// Mitsubishi GX Works2 project: 20国轩1次注液出1031   PLC: Q06UDEH (continued)
  PackCommunication20105 : PackCommunication;
  PackCommunication20106 : PackCommunication;
  PackCommunication20107 : PackCommunication;
  PackCommunication20108 : PackCommunication;
  PackCommunication20109 : PackCommunication;
  PackCommunicationIO20102 : PackCommunicationIO;
  PackCommunicationIO20103 : PackCommunicationIO;
  PackCommunicationIO20104 : PackCommunicationIO;
  PackCommunicationIO20105 : PackCommunicationIO;
  PackCommunicationIO20106 : PackCommunicationIO;
  PackCommunicationIO20107 : PackCommunicationIO;
  PackCommunicationIO20108 : PackCommunicationIO;
  PackCommunicationIO20109 : PackCommunicationIO;
  m_TPU1TaskComplete : TP;  (* U1完成延时 *)
  m_tU1TaskComplete : TIME;  (* U1完成延时 *)
  m_xU1TaskComplete : BOOL;  (* U1完成延时 *)
  m_TPU2TaskComplete : TP;  (* U2完成延时 *)
  m_tU2TaskComplete : TIME;  (* U2完成延时 *)
  m_xU2TaskComplete : BOOL;  (* U2完成延时 *)
  m_TPU3TaskComplete : TP;  (* U3完成延时 *)
  m_tU3TaskComplete : TIME;  (* U3完成延时 *)
  m_xU3TaskComplete : BOOL;  (* U3完成延时 *)
  m_TPU4TaskComplete : TP;  (* U4完成延时 *)
  m_tU4TaskComplete : TIME;  (* U4完成延时 *)
  m_xU4TaskComplete : BOOL;  (* U4完成延时 *)
  m_TonU1TaskStart : TON;  (* U1任务开始延时 *)
  m_tU1TaskStart : TIME;  (* U1任务开始延时 *)
  m_xU1TaskStart : BOOL;  (* U1任务开始延时 *)
  m_TonU2TaskStart : TON;  (* U2任务开始延时 *)
  m_tU2TaskStart : TIME;  (* U2任务开始延时 *)
  m_xU2TaskStart : BOOL;  (* U2任务开始延时 *)
  m_TonU3TaskStart : TON;  (* U3任务开始延时 *)
  m_tU3TaskStart : TIME;  (* U3任务开始延时 *)
  m_xU3TaskStart : BOOL;  (* U3任务开始延时 *)
  m_TonU4TaskStart : TON;  (* U4任务开始延时 *)
  m_tU4TaskStart : TIME;  (* U4任务开始延时 *)
  m_xU4TaskStart : BOOL;  (* U4任务开始延时 *)
  ConveyorIO201221 : ConveyorIO;  (* 虚构的 *)
  Conveyor201221 : Conveyor;  (* 虚构的 *)
  ConveyorIO20119 : ConveyorIO;
  Conveyor20119 : Conveyor;
END_VAR
Conveyor20101(ConveyorMotor:=	ConveyorIO20101);	
(*ConveyorIO20101.xPosLimit:=XA; 	*)
(*ConveyorIO20101.xNegLimit:=X7F; 	*)
ConveyorIO20101.xCWPresent:=X8; 
ConveyorIO20101.xNegLimit:=NOT X9;
(*ConveyorIO20101.xCCWPresent:=X9; 	*)
Y208:=ConveyorIO20101.xMotorCW; 	
Y209:=ConveyorIO20101.xMotorCCW; 	
ConveyorIO20101.xForward:=M500; 	
ConveyorIO20101.xBackward:=M501; 	
M301:= NOT ConveyorIO20101.xEmpty; 	
F401:=ConveyorIO20101.xError; 	
ConveyorIO20101.diDeviceID:=20101; 
ConveyorIO20101.tLoadDelay:=T#2s;	

Conveyor20102(ConveyorMotor:=	ConveyorIO20102);
ConveyorIO20102.xCCWPresent:=X13; 	
Y20A:=ConveyorIO20102.xMotorCW; 	
Y20B:=ConveyorIO20102.xMotorCCW; 	
ConveyorIO20102.xForward:=M502; 	
ConveyorIO20102.xBackward:=M503; 	
M302:= NOT ConveyorIO20102.xEmpty; 	
F402:=ConveyorIO20102.xError; 	
ConveyorIO20102.diDeviceID:=20102;
ConveyorIO20102.tLoadDelay:=T#7s; 
ConveyorIO20102.xloadCCW:=1;	

Conveyor201021(ConveyorMotor:=	ConveyorIO201021);	
ConveyorIO201021.xCWPresent:=X76; 	
M334:= NOT ConveyorIO201021.xEmpty; 	
F434:=ConveyorIO201021.xError; 	
ConveyorIO201021.diDeviceID:=20102; 	
ConveyorIO201021.tLoadDelay:=T#2s;

Conveyor20103(ConveyorMotor:=	ConveyorIO20103);	
ConveyorIO20103.xCCWPresent:=X14; 	
Y20C:=ConveyorIO20103.xMotorCW; 	
Y20D:=ConveyorIO20103.xMotorCCW; 	
ConveyorIO20103.xForward:=M504; 	
ConveyorIO20103.xBackward:=M505; 	
M303:= NOT ConveyorIO20103.xEmpty; 	
F403:=ConveyorIO20103.xError; 	
ConveyorIO20103.diDeviceID:=20103; 
ConveyorIO20103.tLoadDelay:=T#7s; 	
ConveyorIO20103.xloadCCW:=1;	

Conveyor201031(ConveyorMotor:=	ConveyorIO201031);	
ConveyorIO201031.xCWPresent:=X77; 	
M335:= NOT ConveyorIO201031.xEmpty; 	
F435:=ConveyorIO201031.xError; 	
ConveyorIO201031.diDeviceID:=20103; 	
ConveyorIO201031.tLoadDelay:=T#2s;

Conveyor20104(ConveyorMotor:=	ConveyorIO20104);	
ConveyorIO20104.xCCWPresent:=X15; 	
Y20E:=ConveyorIO20104.xMotorCW; 	
Y20F:=ConveyorIO20104.xMotorCCW; 	
ConveyorIO20104.xForward:=M506; 	
ConveyorIO20104.xBackward:=M507; 	
M304:= NOT ConveyorIO20104.xEmpty; 	
F404:=ConveyorIO20104.xError; 	
ConveyorIO20104.diDeviceID:=20104; 
ConveyorIO20104.tLoadDelay:=T#7s; 	
ConveyorIO20104.xloadCCW:=1;		


Conveyor201041(ConveyorMotor:=	ConveyorIO201041);	
ConveyorIO201041.xCWPresent:=X78; 	
M336:= NOT ConveyorIO201041.xEmpty; 	
F436:=ConveyorIO201041.xError; 	
ConveyorIO201041.diDeviceID:=20104; 	
ConveyorIO201041.tLoadDelay:=T#2s;

Conveyor20105(ConveyorMotor:=	ConveyorIO20105);	
ConveyorIO20105.xCCWPresent:=X16; 	
Y210:=ConveyorIO20105.xMotorCW; 	
Y211:=ConveyorIO20105.xMotorCCW; 	
ConveyorIO20105.xForward:=M508; 	
ConveyorIO20105.xBackward:=M509; 	
M305:= NOT ConveyorIO20105.xEmpty; 	
F405:=ConveyorIO20105.xError; 	
ConveyorIO20105.diDeviceID:=20105;		
ConveyorIO20105.tLoadDelay:=T#7s; 	
ConveyorIO20105.xloadCCW:=1;	
				
Conveyor201051(ConveyorMotor:=	ConveyorIO201051);	
ConveyorIO201051.xCWPresent:=X79; 	
M337:= NOT ConveyorIO201051.xEmpty; 	
F437:=ConveyorIO201051.xError; 	
ConveyorIO201051.diDeviceID:=20105; 	
ConveyorIO201051.tLoadDelay:=T#2s;

Conveyor20106(ConveyorMotor:=	ConveyorIO20106);	(*电池X9C*)
ConveyorIO20106.xCCWPresent:=X18; 	
Y212:=ConveyorIO20106.xMotorCW; 	
Y213:=ConveyorIO20106.xMotorCCW; 	
ConveyorIO20106.xForward:=M510; 	
ConveyorIO20106.xBackward:=M511; 	
M306:= NOT ConveyorIO20106.xEmpty; 	
F406:=ConveyorIO20106.xError; 	
ConveyorIO20106.diDeviceID:=20106; 
ConveyorIO20106.tLoadDelay:=T#7s;
ConveyorIO20106.xloadCCW:=1;	 		

Conveyor201061(ConveyorMotor:=	ConveyorIO201061);	
ConveyorIO201061.xCWPresent:=X7A; 	
M338:= NOT ConveyorIO201061.xEmpty; 	
F438:=ConveyorIO201061.xError; 	
ConveyorIO201061.diDeviceID:=20106;
ConveyorIO201061.tLoadDelay:=T#2s; 	

Conveyor20107(ConveyorMotor:=	ConveyorIO20107);	(*电池X9D*)
ConveyorIO20107.xCCWPresent:=X19; 	
Y214:=ConveyorIO20107.xMotorCW; 	
Y215:=ConveyorIO20107.xMotorCCW; 	
ConveyorIO20107.xForward:=M512; 	
ConveyorIO20107.xBackward:=M513; 	
M307:= NOT ConveyorIO20107.xEmpty; 	
F407:=ConveyorIO20107.xError; 	
ConveyorIO20107.diDeviceID:=20107; 
ConveyorIO20107.tLoadDelay:=T#7s; 	
ConveyorIO20107.xloadCCW:=1;	

Conveyor201071(ConveyorMotor:=	ConveyorIO201071);	
ConveyorIO201071.xCWPresent:=X7B; 	
M339:= NOT ConveyorIO201071.xEmpty; 	
F439:=ConveyorIO201071.xError; 	
ConveyorIO201071.diDeviceID:=20107; 	
ConveyorIO201071.tLoadDelay:=T#2s;

Conveyor20108(ConveyorMotor:=	ConveyorIO20108);	(*电池x9e*)
ConveyorIO20108.xCCWPresent:=X1A; 	
Y216:=ConveyorIO20108.xMotorCW; 	
Y217:=ConveyorIO20108.xMotorCCW; 	
ConveyorIO20108.xForward:=M514; 	
ConveyorIO20108.xBackward:=M515; 	
M308:= NOT ConveyorIO20108.xEmpty; 	
F408:=ConveyorIO20108.xError; 	
ConveyorIO20108.diDeviceID:=20108; 
ConveyorIO20108.tLoadDelay:=T#7s; 
ConveyorIO20108.xloadCCW:=1;			

Conveyor201081(ConveyorMotor:=	ConveyorIO201081);	
ConveyorIO201081.xCWPresent:=X7C; 	
M340:= NOT ConveyorIO201081.xEmpty; 	
F440:=ConveyorIO201081.xError; 	
ConveyorIO201081.diDeviceID:=20108; 	
ConveyorIO201081.tLoadDelay:=T#2s;


Conveyor20109(ConveyorMotor:=	ConveyorIO20109);	
ConveyorIO20109.xCCWPresent:=X1B; 	
Y218:=ConveyorIO20109.xMotorCW; 	
Y219:=ConveyorIO20109.xMotorCCW; 	
ConveyorIO20109.xForward:=M516; 	
ConveyorIO20109.xBackward:=M517; 	
M309:= NOT ConveyorIO20109.xEmpty; 	
F409:=ConveyorIO20109.xError; 	
ConveyorIO20109.diDeviceID:=20109;
ConveyorIO20109.tLoadDelay:=T#7s; 	 
ConveyorIO20109.xloadCCW:=1;		
(*电池检测X9F*)

Conveyor201091(ConveyorMotor:=	ConveyorIO201091);	
ConveyorIO201091.xCWPresent:=X7D; 	
M341:= NOT ConveyorIO201091.xEmpty; 	
F441:=ConveyorIO201091.xError; 	
ConveyorIO201091.diDeviceID:=20109;		
ConveyorIO201091.tLoadDelay:=T#2s;

Conveyor20110(ConveyorMotor:=	ConveyorIO20110);	
Y21A:=ConveyorIO20110.xMotorCW; 	
ConveyorIO20110.xForward:=M518; 	
M310:= NOT ConveyorIO20110.xEmpty; 	
F410:=ConveyorIO20110.xError; 	
ConveyorIO20110.diDeviceID:=20110; 
ConveyorIO20110.tLoadDelay:=T#5s;	
ConveyorIO20110.tUnloadAlarmDelay:=T#40s;

Conveyor20111(ConveyorMotor:=	ConveyorIO20111);	
Y21B:=ConveyorIO20111.xMotorCW; 	
ConveyorIO20111.xForward:=M519; 	
M311:= NOT ConveyorIO20111.xEmpty; 	
F411:=ConveyorIO20111.xError; 	
ConveyorIO20111.diDeviceID:=20111;
ConveyorIO20111.tLoadDelay:=T#4s;	 	

Conveyor20112(ConveyorMotor:=	ConveyorIO20112);	
ConveyorIO20112.xCWPresent:=X17; (*暂时改为XE，调试用。实际X17*)	
Y21C:=ConveyorIO20112.xMotorCW; 	
ConveyorIO20112.xForward:=M520; 	
M312:= NOT ConveyorIO20112.xEmpty; 	
F412:=ConveyorIO20112.xError; 	
ConveyorIO20112.diDeviceID:=20112; 	

Conveyor20113(ConveyorMotor:=	ConveyorIO20113);	
Y21D:=ConveyorIO20113.xMotorCW; 	
ConveyorIO20113.xForward:=M521; 	
M313:= NOT ConveyorIO20113.xEmpty; 	
F413:=ConveyorIO20113.xError; 	
ConveyorIO20113.diDeviceID:=20113;
ConveyorIO20113.tLoadDelay:=T#4s;	 	

Conveyor20114(ConveyorMotor:=	ConveyorIO20114);	
Y21E:=ConveyorIO20114.xMotorCW; 	
ConveyorIO20114.xForward:=M522; 	
M314:= NOT ConveyorIO20114.xEmpty; 	
F414:=ConveyorIO20114.xError; 	
ConveyorIO20114.diDeviceID:=20114; 	
ConveyorIO20114.tLoadDelay:=T#4s;	
ConveyorIO20114.tUnloadAlarmDelay:=T#40s;


Conveyor20115(ConveyorMotor:=	ConveyorIO20115);	
ConveyorIO20115.xCWPresent:=X1C; 
M315:= NOT ConveyorIO20116.xEmpty; 	
F415:=ConveyorIO20116.xError; 		
ConveyorIO20115.diDeviceID:=20115;	
ConveyorIo20115.tLoadDelay:=T#4500ms;	

Conveyor20116(ConveyorMotor:=	ConveyorIO20116);	
ConveyorIO20116.xCWPresent:=X1C; 	
Y21F:=ConveyorIO20116.xMotorCW; 	
ConveyorIO20116.xForward:=M523; 	
M316:= NOT ConveyorIO20116.xEmpty; 	
F416:=ConveyorIO20116.xError; 	
ConveyorIO20116.diDeviceID:=20116; 	

Conveyor20117(ConveyorMotor:=	ConveyorIO20117);	
ConveyorIO20117.xCWPresent:=X1E; 	
Y220:=ConveyorIO20117.xMotorCW; 	
ConveyorIO20117.xForward:=M524; 	
M317:= NOT ConveyorIO20117.xEmpty; 	
F417:=ConveyorIO20117.xError; 	
ConveyorIO20117.diDeviceID:=20117; 	

Conveyor20118(ConveyorMotor:=	ConveyorIO20118);	
ConveyorIO20118.xCWPresent:=X1F; 	
Y221:=ConveyorIO20118.xMotorCW; 	
ConveyorIO20118.xForward:=M525; 	
M318:= NOT ConveyorIO20118.xEmpty; 	
F418:=ConveyorIO20118.xError; 	
ConveyorIO20118.diDeviceID:=20118; 	

Conveyor20119(ConveyorMotor:=	ConveyorIO20119);	
ConveyorIO20119.xCWPresent:=X20; 	
Y222:=ConveyorIO20119.xMotorCW;	
ConveyorIO20119.xForward:=M526; 	
M319:= NOT ConveyorIO20119.xEmpty; 	
F419:=ConveyorIO20119.xError; 	
ConveyorIO20119.diDeviceID:=20119; 	

Conveyor201191(ConveyorMotor:= ConveyorIO201191 );
ConveyorIO201191 .xCWPresent:=X20;
ConveyorIO201191 .diDeviceID:=201191;

Conveyor20122(ConveyorMotor:=	ConveyorIO20122);	
ConveyorIO20122.xCWPresent:=X23;
Y226:=ConveyorIO20122.xMotorCW; 	
ConveyorIO20122.xForward:=M530; 	
M322:= NOT ConveyorIO20122.xEmpty; 	
F422:=ConveyorIO20122.xError; 	
ConveyorIO20122.diDeviceID:=20122; 	

Conveyor201221(ConveyorMotor:= ConveyorIO201221 );
ConveyorIO201221 .xCWPresent:=X23;
ConveyorIO201221 .diDeviceID:=201221;
ConveyorIO201221.tLoadDelay:=T#6s;

Conveyor20123(ConveyorMotor:=	ConveyorIO20123);	
ConveyorIO20123.xCWPresent:=X25; 	
Y227:=ConveyorIO20123.xMotorCW; 	
ConveyorIO20123.xForward:=M531; 	
M323:= NOT ConveyorIO20123.xEmpty; 	
F423:=ConveyorIO20123.xError; 	
ConveyorIO20123.diDeviceID:=20123; 	

Conveyor20124(ConveyorMotor:=	ConveyorIO20124);	
ConveyorIO20124.xCWPresent:=X26; 	
Y228:=ConveyorIO20124.xMotorCW; 	
ConveyorIO20124.xForward:=M532; 	
M324:= NOT ConveyorIO20124.xEmpty; 	
F424:=ConveyorIO20124.xError; 	
ConveyorIO20124.diDeviceID:=20124; 	

Conveyor20125(ConveyorMotor:=	ConveyorIO20125);	
ConveyorIO20125.xCWPresent:=X27; 	
Y225:=ConveyorIO20125.xMotorCW; 	
ConveyorIO20125.xForward:=M533; 	
M325:= NOT ConveyorIO20125.xEmpty; 	
F425:=ConveyorIO20125.xError; 	
ConveyorIO20125.diDeviceID:=20125;
ConveyorIO20125.tLoadDelay:=T#6s; 	

Conveyor20126(ConveyorMotor:=	ConveyorIO20126);	
ConveyorIO20126.xCWPresent:=X27; 	
Y224:=ConveyorIO20126.xMotorCW; 	
ConveyorIO20126.xForward:=M534; 	
M326:= NOT ConveyorIO20126.xEmpty; 	
F426:=ConveyorIO20126.xError; 	
ConveyorIO20126.diDeviceID:=20126; 	

Conveyor20127(ConveyorMotor:=	ConveyorIO20127);	
ConveyorIO20127.xCWPresent:=X29; 	
Y223:=ConveyorIO20127.xMotorCW; 	
ConveyorIO20127.xForward:=M535; 	
M327:= NOT ConveyorIO20127.xEmpty; 	
F427:=ConveyorIO20127.xError; 	
ConveyorIO20127.diDeviceID:=20127; 	

Conveyor20128(ConveyorMotor:=	ConveyorIO20128);	
ConveyorIO20128.xCWPresent:=X2A; 	(*暂时改为XF，调试用，X2A*)
Y22A:=ConveyorIO20128.xMotorCW; 	
ConveyorIO20128.xForward:=M536; 	
M328:= NOT ConveyorIO20128.xEmpty; 	
F428:=ConveyorIO20128.xError; 	
ConveyorIO20128.diDeviceID:=20128; 	

Conveyor20129(ConveyorMotor:=	ConveyorIO20129);	
ConveyorIO20129.xCWPresent:=X2B; 	
Y22D:=ConveyorIO20129.xMotorCW; 	
ConveyorIO20129.xForward:=M537; 	
M329:= NOT ConveyorIO20129.xEmpty; 	
F429:=ConveyorIO20129.xError; 	
ConveyorIO20129.diDeviceID:=20129; 	

Conveyor20130(ConveyorMotor:=	ConveyorIO20130);	
ConveyorIO20130.xPosLimit:= NOT X70; 	
ConveyorIO20130.xCWPresent:=X2C; 	
Y22E:=ConveyorIO20130.xMotorCW; 	
ConveyorIO20130.xForward:=M538; 	
M330:= NOT ConveyorIO20130.xEmpty; 	
F430:=ConveyorIO20130.xError; 	
ConveyorIO20130.diDeviceID:=20130; 	
			
UConveyor20301(	ConveyorIOLeft:= ConveyorIO20102,
 				ConveyorIORight:= ConveyorIO20103,
 				ConveyorIODown:= ConveyorIO20110,
 				UConveyorIO:= UConveyorIO20301);
UConveyorIO20301.xLiftCylinderRetractDetect1:=X30;
UConveyorIO20301.xLiftCylinderExtendDetect1:=X31;
Y236:=UConveyorIO20301.xLiftCylinderExtend1;
Y278:=UConveyorIO20301.xExitBarCylinderRetract1;
UConveyorIO20301.xLiftCylinderRetractDetect2:=X33;
UConveyorIO20301.xLiftCylinderExtendDetect2:=X32;
Y238:=UConveyorIO20301.xLiftCylinderExtend2;
Y279:=UConveyorIO20301.xExitBarCylinderRetract2;
UConveyorIO20301.xLiftCylinderExtendButton1:=M548;
UConveyorIO20301.xExitBarCylinderRetractButton1:=M549;
UConveyorIO20301.xLiftCylinderExtendButton2:=M550;
UConveyorIO20301.xExitBarCylinderRetractButton2:=M551;
F448:=UConveyorIO20301.xOvertimeAlarm ;
UConveyorIO20301.xBatteryDetect1:=0(*X98*);
UConveyorIO20301.xBatteryDetect2:=0(*X99*);

UConveyor20303(	ConveyorIOLeft:= ConveyorIO20104,	
 				ConveyorIORight:= ConveyorIO20105,	
 				ConveyorIODown:= ConveyorIO20111,	
 				UConveyorIO:= UConveyorIO20303);
UConveyorIO20303.xLiftCylinderRetractDetect1:=X35;
UConveyorIO20303.xLiftCylinderExtendDetect1:=X34;
Y23A:=UConveyorIO20303.xLiftCylinderExtend1;
Y27A:=UConveyorIO20303.xExitBarCylinderRetract1;
UConveyorIO20303.xLiftCylinderRetractDetect2:=X37;
UConveyorIO20303.xLiftCylinderExtendDetect2:=X36;
Y23C:=UConveyorIO20303.xLiftCylinderExtend2;
Y27B:=UConveyorIO20303.xExitBarCylinderRetract2;
UConveyorIO20303.xLiftCylinderExtendButton1:=M552;
UConveyorIO20303.xExitBarCylinderRetractButton1:=M553;
UConveyorIO20303.xLiftCylinderExtendButton2:=M554;
UConveyorIO20303.xExitBarCylinderRetractButton2:=M555;
F449:=UConveyorIO20303.xOvertimeAlarm ;
UConveyorIO20303.xBatteryDetect1:=0(*X9A*);
UConveyorIO20303.xBatteryDetect2:=0(*X9B*);

UConveyor20305(	ConveyorIOLeft:= ConveyorIO20106,	
 				ConveyorIORight:= ConveyorIO20107,	
 				ConveyorIODown:= ConveyorIO20113,
 				UConveyorIO:= UConveyorIO20305);
UConveyorIO20305.xLiftCylinderRetractDetect1:=X39;
UConveyorIO20305.xLiftCylinderExtendDetect1:=X38;
Y23E:=UConveyorIO20305.xLiftCylinderExtend1;
Y27C:=UConveyorIO20305.xExitBarCylinderRetract1;
UConveyorIO20305.xLiftCylinderRetractDetect2:=X3B;
UConveyorIO20305.xLiftCylinderExtendDetect2:=X3A;
Y240:=UConveyorIO20305.xLiftCylinderExtend2;
Y27D:=UConveyorIO20305.xExitBarCylinderRetract2;
UConveyorIO20305.xLiftCylinderExtendButton1:=M556;
UConveyorIO20305.xExitBarCylinderRetractButton1:=M557;
UConveyorIO20305.xLiftCylinderExtendButton2:=M558;
UConveyorIO20305.xExitBarCylinderRetractButton2:=M559;
F450:=UConveyorIO20305.xOvertimeAlarm ;
UConveyorIO20305.xBatteryDetect1:=0(*X9C*);
UConveyorIO20305.xBatteryDetect2:=0(*X9D*);

UConveyor20307(	ConveyorIOLeft:= ConveyorIO20109,	
 				ConveyorIORight:= ConveyorIO20108,	
 				ConveyorIODown:= ConveyorIO20114,	
 				UConveyorIO:= UConveyorIO20307);
UConveyorIO20307.xLiftCylinderRetractDetect1:=X3F;
UConveyorIO20307.xLiftCylinderExtendDetect1:=X3E;
Y244:=UConveyorIO20307.xLiftCylinderExtend1;
Y27E:=UConveyorIO20307.xExitBarCylinderRetract1;
UConveyorIO20307.xLiftCylinderRetractDetect2:=X3D;
UConveyorIO20307.xLiftCylinderExtendDetect2:=X3C;
Y242:=UConveyorIO20307.xLiftCylinderExtend2;
Y27F:=UConveyorIO20307.xExitBarCylinderRetract2;
UConveyorIO20307.xLiftCylinderExtendButton1:=M560;
UConveyorIO20307.xExitBarCylinderRetractButton1:=M561;
UConveyorIO20307.xLiftCylinderExtendButton2:=M562;
UConveyorIO20307.xExitBarCylinderRetractButton2:=M563;
F451:=UConveyorIO20307.xOvertimeAlarm ;
UConveyorIO20307.xBatteryDetect1:=0;(*X9E;*)
UConveyorIO20307.xBatteryDetect2:=0;(*X9F;*)
(*U型结构出口处的夹紧气缸*)
Y254:=m_xCatchCylinder[2];
Y256:=m_xCatchCylinder[3];
Y258:=m_xCatchCylinder[4];
Y25A:=m_xCatchCylinder[5];
Y25E:=m_xCatchCylinder[6];
Y25C:=m_xCatchCylinder[7];
Y260:=m_xCatchCylinder[8];
Y262:=m_xCatchCylinder[9];
Switch20309(	ConveyorEntryIO:= ConveyorIO20115,	
 		ConveyorExitIO:=ConveyorIO20116,	
 		SwitchIO:=SwitchIO20309);
SwitchIO20309.xLiftCylinderRetractDetect:=X41;				
SwitchIO20309.xLiftCylinderExtendDetect:=X40;				
Y246:=SwitchIO20309.xLiftCylinderExtend;				
SwitchIO20309.xLiftCylinderExtendButton:=M544;
SwitchIO20309.xLiftCylinderRetractButton:=NOT M544;
F444:=SwitchIO20309.xOvertimeAlarm ;				

Switch20310(	ConveyorEntryIO:= ConveyorIO20119,	
 		ConveyorExitIO:=ConveyorIO201191,	
 		SwitchIO:=SwitchIO20310);
SwitchIO20310.xLiftCylinderRetractDetect:=X43;				
SwitchIO20310.xLiftCylinderExtendDetect:=X42;				
Y248:=SwitchIO20310.xLiftCylinderExtend;				
SwitchIO20310.xLiftCylinderExtendButton:=M545;	
SwitchIO20310.xLiftCylinderRetractButton:=NOT M545;				
F445:=SwitchIO20310.xOvertimeAlarm ;				

Switch20311(	ConveyorEntryIO:= ConveyorIO201221,	
 		ConveyorExitIO:=ConveyorIO20122,	
 		SwitchIO:=SwitchIO20311);
SwitchIO20311.xLiftCylinderRetractDetect:=X45;				
SwitchIO20311.xLiftCylinderExtendDetect:=X44;				
Y24A:=SwitchIO20311.xLiftCylinderExtend;				
SwitchIO20311.xLiftCylinderExtendButton:=M546;	
SwitchIO20311.xLiftCylinderRetractButton:=NOT M546;				
F446:=SwitchIO20311.xOvertimeAlarm ;				

Switch20312(	ConveyorEntryIO:= ConveyorIO20125,	
 		ConveyorExitIO:=ConveyorIO20126,	
 		SwitchIO:=SwitchIO20312);
SwitchIO20312.xLiftCylinderRetractDetect:=X47;				
SwitchIO20312.xLiftCylinderExtendDetect:=X46;				
Y24C:=SwitchIO20312.xLiftCylinderExtend;				
SwitchIO20312.xLiftCylinderExtendButton:=M547;
SwitchIO20312.xLiftCylinderRetractButton:=NOT M547;				
F447:=SwitchIO20312.xOvertimeAlarm ;				

Lifter20201(ShuttleCarInOut:=LifterIO20201);
LifterIO20201.xCylinder:=1;
Y235:=LifterIO20201.xCW;
Y234:=LifterIO20201.xCCW;
LifterIO20201.xForward:=M542;
LifterIO20201.xBackward:=M543;
ShuttleCarCurrentPosition(X2F OR X2E,X2E,X2F,FALSE,LifterIO20201.iCurrentPos);
F443:=LifterIO20201.xOvertimeAlarm ;
LifterIO20201.diDeviceID:=20201;

Robot20901(FanucRobotIO:=RobotIO20901);
Robot20902(FanucRobotIO:=RobotIO20902);
Robot20903(FanucRobotIO:=RobotIO20903);
Robot20904(FanucRobotIO:=RobotIO20904);

	PackCommunication20102(ConveyorIO:=ConveyorIO201021,
 	PackCommunicationIO:=PackCommunicationIO20102 ,
 	FanucRobotIO:= RobotIO20901 ,
 	i_arrxPresentDetect:=g_xRobot1BatteryDetect);
	PackCommunicationIO20102.i_iResponsPCPLC:=D2001;
	PackCommunicationIO20102.i_iPackDoneAknPCPLC:=D2002;
	PackCommunicationIO20102.i_iSinglePackResponsePCPLC:=D2003;
	PackCommunicationIO20102.i_iSinglePackDoneAknPCPLC:=D2004;
	D3001:=PackCommunicationIO20102.o_iRequestPLCPC;
	D3002:=PackCommunicationIO20102.o_iPackDonePLCPC;
	D3003:=PackCommunicationIO20102.o_iSinglePackRequestPLCPC;
	D3004:=PackCommunicationIO20102.o_iSinglePackDonePLCPC;
	D3005:=PackCommunicationIO20102.o_iXCoordinatePLCPC;
	D3006:=PackCommunicationIO20102.o_iYCoordinatePLCPC;(*?
	FOR Z0:=0 TO 120 BY 1 DO(*120是因为15*8，15个字存一个码，8是因为一排有8个电池*)(*?
		D3007Z0:=PackCommunicationIO20102.o_arrwCode[DIV( Z0 , 8 )].arrwCode[ Z0 MOD 8 ];
	END_FOR;?*)
		
	PackCommunication20103(ConveyorIO:=ConveyorIO201031,
 	PackCommunicationIO:=PackCommunicationIO20103 ,
 	FanucRobotIO:= RobotIO20901 ,
 	i_arrxPresentDetect:=g_xRobot1BatteryDetect);
	PackCommunicationIO20103.i_iResponsPCPLC:=D2011;
	PackCommunicationIO20103.i_iPackDoneAknPCPLC:=D2012;
	PackCommunicationIO20103.i_iSinglePackResponsePCPLC:=D2013;
	PackCommunicationIO20103.i_iSinglePackDoneAknPCPLC:=D2014;
	D3201:=PackCommunicationIO20103.o_iRequestPLCPC;
	D3202:=PackCommunicationIO20103.o_iPackDonePLCPC;
	D3203:=PackCommunicationIO20103.o_iSinglePackRequestPLCPC;
	D3204:=PackCommunicationIO20103.o_iSinglePackDonePLCPC;
	D3205:=PackCommunicationIO20103.o_iXCoordinatePLCPC;
	D3206:=PackCommunicationIO20103.o_iYCoordinatePLCPC;(*?
	FOR Z0:=0 TO 120 BY 1 DO
		D3207Z0:=PackCommunicationIO20103.o_arrwCode[DIV( Z0 , 8 )].arrwCode[ Z0 MOD 8 ];
	END_FOR;?*)
	
	PackCommunication20104(ConveyorIO:=ConveyorIO201041,
 	PackCommunicationIO:=PackCommunicationIO20104 ,
 	FanucRobotIO:= RobotIO20902 ,
 	i_arrxPresentDetect:=g_xRobot2BatteryDetect);
	PackCommunicationIO20104.i_iResponsPCPLC:=D2021;
	PackCommunicationIO20104.i_iPackDoneAknPCPLC:=D2022;
	PackCommunicationIO20104.i_iSinglePackResponsePCPLC:=D2023;
	PackCommunicationIO20104.i_iSinglePackDoneAknPCPLC:=D2024;
	D3401:=PackCommunicationIO20104.o_iRequestPLCPC;
	D3402:=PackCommunicationIO20104.o_iPackDonePLCPC;
	D3403:=PackCommunicationIO20104.o_iSinglePackRequestPLCPC;
	D3404:=PackCommunicationIO20104.o_iSinglePackDonePLCPC;
	D3405:=PackCommunicationIO20104.o_iXCoordinatePLCPC;
	D3406:=PackCommunicationIO20104.o_iYCoordinatePLCPC;(*?
	FOR Z0:=0 TO 120 BY 1 DO
		D3407Z0:=PackCommunicationIO20104.o_arrwCode[DIV( Z0 , 8 )].arrwCode[ Z0 MOD 8 ];
	END_FOR;?*)
	
	PackCommunication20105(ConveyorIO:=ConveyorIO201051,
 	PackCommunicationIO:=PackCommunicationIO20105 ,
 	FanucRobotIO:= RobotIO20902 ,
 	i_arrxPresentDetect:=g_xRobot2BatteryDetect);
	PackCommunicationIO20105.i_iResponsPCPLC:=D2031;
	PackCommunicationIO20105.i_iPackDoneAknPCPLC:=D2032;
	PackCommunicationIO20105.i_iSinglePackResponsePCPLC:=D2033;
	PackCommunicationIO20105.i_iSinglePackDoneAknPCPLC:=D2034;
	D3601:=PackCommunicationIO20105.o_iRequestPLCPC;
	D3602:=PackCommunicationIO20105.o_iPackDonePLCPC;
	D3603:=PackCommunicationIO20105.o_iSinglePackRequestPLCPC;
	D3604:=PackCommunicationIO20105.o_iSinglePackDonePLCPC;
	D3605:=PackCommunicationIO20105.o_iXCoordinatePLCPC;
	D3606:=PackCommunicationIO20105.o_iYCoordinatePLCPC;(*?
	FOR Z0:=0 TO 120 BY 1 DO
		D3607Z0:=PackCommunicationIO20105.o_arrwCode[DIV( Z0 , 8 )].arrwCode[ Z0 MOD 8 ];
	END_FOR;?*)
	
	PackCommunication20106(ConveyorIO:=ConveyorIO201061,
 	PackCommunicationIO:=PackCommunicationIO20106 ,
 	FanucRobotIO:= RobotIO20903 ,
 	i_arrxPresentDetect:=g_xRobot3BatteryDetect);
	PackCommunicationIO20106.i_iResponsPCPLC:=D2041;
	PackCommunicationIO20106.i_iPackDoneAknPCPLC:=D2042;
	PackCommunicationIO20106.i_iSinglePackResponsePCPLC:=D2043;
	PackCommunicationIO20106.i_iSinglePackDoneAknPCPLC:=D2044;
	D3801:=PackCommunicationIO20106.o_iRequestPLCPC;
	D3802:=PackCommunicationIO20106.o_iPackDonePLCPC;
	D3803:=PackCommunicationIO20106.o_iSinglePackRequestPLCPC;
	D3804:=PackCommunicationIO20106.o_iSinglePackDonePLCPC;
	D3805:=PackCommunicationIO20106.o_iXCoordinatePLCPC;
	D3806:=PackCommunicationIO20106.o_iYCoordinatePLCPC;(*?
	FOR Z0:=0 TO 120 BY 1 DO
		D3807Z0:=PackCommunicationIO20106.o_arrwCode[DIV( Z0 , 8 )].arrwCode[ Z0 MOD 8 ];
	END_FOR;?*)
	
	PackCommunication20107(ConveyorIO:=ConveyorIO201071,
 	PackCommunicationIO:=PackCommunicationIO20107 ,
 	FanucRobotIO:= RobotIO20903 ,
 	i_arrxPresentDetect:=g_xRobot3BatteryDetect);
	PackCommunicationIO20107.i_iResponsPCPLC:=D2051;
	PackCommunicationIO20107.i_iPackDoneAknPCPLC:=D2052;
	PackCommunicationIO20107.i_iSinglePackResponsePCPLC:=D2053;
	PackCommunicationIO20107.i_iSinglePackDoneAknPCPLC:=D2054;
	D4001:=PackCommunicationIO20107.o_iRequestPLCPC;
	D4002:=PackCommunicationIO20107.o_iPackDonePLCPC;
	D4003:=PackCommunicationIO20107.o_iSinglePackRequestPLCPC;
	D4004:=PackCommunicationIO20107.o_iSinglePackDonePLCPC;
	D4005:=PackCommunicationIO20107.o_iXCoordinatePLCPC;
	D4006:=PackCommunicationIO20107.o_iYCoordinatePLCPC;(*?
	FOR Z0:=0 TO 120 BY 1 DO
		D4007Z0:=PackCommunicationIO20107.o_arrwCode[DIV( Z0 , 8 )].arrwCode[ Z0 MOD 8 ];
	END_FOR;?*)
	
	PackCommunication20108(ConveyorIO:=ConveyorIO201081,
 	PackCommunicationIO:=PackCommunicationIO20108 ,
 	FanucRobotIO:= RobotIO20904 ,
 	i_arrxPresentDetect:=g_xRobot4BatteryDetect);
	PackCommunicationIO20108.i_iResponsPCPLC:=D2061;
	PackCommunicationIO20108.i_iPackDoneAknPCPLC:=D2062;
	PackCommunicationIO20108.i_iSinglePackResponsePCPLC:=D2063;
	PackCommunicationIO20108.i_iSinglePackDoneAknPCPLC:=D2064;
	D4201:=PackCommunicationIO20108.o_iRequestPLCPC;
	D4202:=PackCommunicationIO20108.o_iPackDonePLCPC;
	D4203:=PackCommunicationIO20108.o_iSinglePackRequestPLCPC;
	D4204:=PackCommunicationIO20108.o_iSinglePackDonePLCPC;
	D4205:=PackCommunicationIO20108.o_iXCoordinatePLCPC;
	D4206:=PackCommunicationIO20108.o_iYCoordinatePLCPC;(*?
	FOR Z0:=0 TO 120 BY 1 DO
		D4207Z0:=PackCommunicationIO20108.o_arrwCode[DIV( Z0 , 8 )].arrwCode[ Z0 MOD 8 ];
	END_FOR;?*)
	
	PackCommunication20109(ConveyorIO:=ConveyorIO201091,
 	PackCommunicationIO:=PackCommunicationIO20109,
 	FanucRobotIO:= RobotIO20904,
 	i_arrxPresentDetect:=g_xRobot4BatteryDetect);
	PackCommunicationIO20109.i_iResponsPCPLC:=D2071;
	PackCommunicationIO20109.i_iPackDoneAknPCPLC:=D2072;
	PackCommunicationIO20109.i_iSinglePackResponsePCPLC:=D2073;
	PackCommunicationIO20109.i_iSinglePackDoneAknPCPLC:=D2074;
	D4401:=PackCommunicationIO20109.o_iRequestPLCPC;
	D4402:=PackCommunicationIO20109.o_iPackDonePLCPC;
	D4403:=PackCommunicationIO20109.o_iSinglePackRequestPLCPC;
	D4404:=PackCommunicationIO20109.o_iSinglePackDonePLCPC;
	D4405:=PackCommunicationIO20109.o_iXCoordinatePLCPC;
	D4406:=PackCommunicationIO20109.o_iYCoordinatePLCPC;(*?
	FOR Z0:=0 TO 120 BY 1 DO
		D4407Z0:=PackCommunicationIO20109.o_arrwCode[DIV( Z0 , 8 )].arrwCode[ Z0 MOD 8 ];
	END_FOR;?*)
(******************************************上位机通信数据**************************************************)

(******************************************以上是上位机通信***************************************)
(*任务处理*)
(*提升机生成8个入口的排队任务*)
	Conveyor20101Task(	arrxCondition:=Conveyor20101Condition ,
  		xTaskComplete:=LDP(TRUE,ConveyorIO20101.xEmpty) ,
  		arriTaskStack:=g_iLoadTask,
  		xReset:=g_xResetTask1,
  		iPriority:=m_i20101Task);
	Conveyor20101Condition[1].xCondition:=	ConveyorIO201091.xEmpty 	AND m_xLoadPermit[9];
	Conveyor20101Condition[2].xCondition:=	ConveyorIO201081.xEmpty	AND m_xLoadPermit[8];
	Conveyor20101Condition[3].xCondition:=	ConveyorIO201071.xEmpty	AND m_xLoadPermit[7];
	Conveyor20101Condition[4].xCondition:=	ConveyorIO201061.xEmpty	AND m_xLoadPermit[6];
	Conveyor20101Condition[5].xCondition:=	ConveyorIO201051.xEmpty	AND m_xLoadPermit[5];
	Conveyor20101Condition[6].xCondition:=	ConveyorIO201041.xEmpty	AND m_xLoadPermit[4];
	Conveyor20101Condition[7].xCondition:=	ConveyorIO201031.xEmpty	AND m_xLoadPermit[3];
	Conveyor20101Condition[8].xCondition:=	ConveyorIO201021.xEmpty	AND m_xLoadPermit[2];
	m_xLoadPermit[9]:=M59;(*允许信号，由触摸屏给的·*)
	m_xLoadPermit[8]:=M58;
	m_xLoadPermit[7]:=M57;
	m_xLoadPermit[6]:=M56;
	m_xLoadPermit[5]:=M55;
	m_xLoadPermit[4]:=M54;
	m_xLoadPermit[3]:=M53;
	m_xLoadPermit[2]:=M52;
	(*根据任务生成目标地址	*)
	DMOV(m_i20101Task=1,	20109,	ConveyorIO20101.diDesConveyor);
	DMOV(m_i20101Task=2,	20108,	ConveyorIO20101.diDesConveyor);
	DMOV(m_i20101Task=3,	20107,	ConveyorIO20101.diDesConveyor);
	DMOV(m_i20101Task=4,	20106,	ConveyorIO20101.diDesConveyor);
	DMOV(m_i20101Task=5,	20105,	ConveyorIO20101.diDesConveyor);
	DMOV(m_i20101Task=6,	20104,	ConveyorIO20101.diDesConveyor);
	DMOV(m_i20101Task=7,	20103,	ConveyorIO20101.diDesConveyor);
	DMOV(m_i20101Task=8,	20102,	ConveyorIO20101.diDesConveyor);
	
	(*U1任务处理 *)
	m_TPU1TaskComplete(IN:=ConveyorIO20110.xEmpty ,PT:=t#200ms,Q:= m_xU1TaskComplete,ET:= m_tU1TaskComplete );
	(*这里东西运走之后延时200ms再完成任务，这个时间是防止扫描周期的影响，让U型块先复位，再完成任务*)
Task20301(	xCondition:=TaskCondition20301,
 xTaskComplete:=LDF(TRUE,m_xU1TaskComplete),
 xReset:=g_xResetSingle AND g_diDeviceIDSelect=20110,
 iPriority:=UConveyorIO20301.iTask);
	TaskCondition20301[1]:=NOT ConveyorIO20101.xEmpty  AND LifterIO20201.iCurrentPos=2  AND X2F AND m_i20101Task>0;
	TaskCondition20301[2]:=(NOT ConveyorIO201021.xEmpty AND ConveyorIO201021.diDesConveyor=20115) 
												OR(NOT  ConveyorIO20110.xEmpty AND (ConveyorIO20110.diDesConveyor<>20102 OR ConveyorIO20110.diDesConveyor<>20103)) ;
	TaskCondition20301[3]:=(NOT ConveyorIO201031.xEmpty AND ConveyorIO201031.diDesConveyor=20115)
												OR (NOT  ConveyorIO20110.xEmpty AND(ConveyorIO20110.diDesConveyor<>20102 OR ConveyorIO20110.diDesConveyor<>20103));
	(*U2Task	*)
	m_TPU2TaskComplete(IN:=ConveyorIO20111.xEmpty ,PT:=t#200ms,Q:= m_xU2TaskComplete,ET:= m_tU2TaskComplete );
	Task20303(	xCondition:=TaskCondition20303,
 	xTaskComplete:=LDf(TRUE, m_xU2TaskComplete),
 	xReset:=g_xResetSingle AND g_diDeviceIDSelect=20111,
 	iPriority:=UConveyorIO20303.iTask);
		TaskCondition20303[1]:=NOT ConveyorIO20110.xEmpty AND NOT  (ConveyorIO20110.diDesConveyor=20103 
																OR ConveyorIO20110.diDesConveyor=20102
																OR ConveyorIO20110.diDesConveyor=0)(*不去左，不去右，也不是0，就认为可以接料*);
		TaskCondition20303[2]:=(NOT ConveyorIO201041.xEmpty  AND ConveyorIO201041.diDesConveyor=20115) 
													OR (NOT ConveyorIO20111.xEmpty AND (ConveyorIO20111.diDesConveyor<>20103 OR ConveyorIO20111.diDesConveyor<>20102) );
		TaskCondition20303[3]:=(NOT ConveyorIO201051.xEmpty  AND ConveyorIO201051.diDesConveyor=20115) 
													OR (NOT ConveyorIO20111.xEmpty AND (ConveyorIO20111.diDesConveyor<>20103 OR ConveyorIO20111.diDesConveyor<>20102));
	(*//U3Task*)
	m_TPU3TaskComplete(IN:=ConveyorIO20113.xEmpty ,PT:=t#200ms,Q:= m_xU3TaskComplete,ET:= m_tU3TaskComplete );
	Task20305(	xCondition:=TaskCondition20305,
 	xTaskComplete:=LDF(TRUE,m_xU3TaskComplete),
 	xReset:=g_xResetSingle AND g_diDeviceIDSelect=20113,
 	iPriority:=UConveyorIO20305.iTask);
		TaskCondition20305[1]:=NOT ConveyorIO20112.xEmpty(* AND  (ConveyorIO20112.diDesConveyor=20104 
																OR ConveyorIO20112.diDesConveyor=20105
																OR ConveyorIO20112.diDesConveyor=0);(*不去左，不去右，也不是0，就认为可以接料*) ;
		TaskCondition20305[2]:=(NOT ConveyorIO201061.xEmpty AND ConveyorIO201061.diDesConveyor=20115) 
													OR (NOT ConveyorIO20113.xEmpty AND (ConveyorIO20113.diDesConveyor<>20104 OR ConveyorIO20113.diDesConveyor<>20105));
		TaskCondition20305[3]:=(NOT ConveyorIO201071.xEmpty AND ConveyorIO201071.diDesConveyor=20115)
													OR (NOT ConveyorIO20113.xEmpty AND  (ConveyorIO20113.diDesConveyor<>20104 OR ConveyorIO20113.diDesConveyor<>20105));
	(*//U4Task*)
	m_TPU4TaskComplete(IN:=ConveyorIO20114.xEmpty ,PT:=t#200ms,Q:= m_xU4TaskComplete,ET:= m_tU4TaskComplete );
	Task20307(	xCondition:=TaskCondition20307,
 	xTaskComplete:=LDF(TRUE, m_xU4TaskComplete),
 	xReset:=g_xResetSingle AND g_diDeviceIDSelect=20114,
 	iPriority:=UConveyorIO20307.iTask);
		TaskCondition20307[1]:=NOT ConveyorIO20113.xEmpty  AND NOT (ConveyorIO20113.diDesConveyor=20109
																OR ConveyorIO20113.diDesConveyor=20108
																OR ConveyorIO20113.diDesConveyor=0)
																AND ConveyorIo20115.xEmpty;		
		TaskCondition20307[2]:=((NOT ConveyorIO201091.xEmpty AND ConveyorIO201091.diDesConveyor=20115)
													OR (NOT ConveyorIO20114.xEmpty AND (ConveyorIO20114.diDesConveyor<>20109 OR ConveyorIO20114.diDesConveyor<>20108) ))
													AND ConveyorIo20115.xEmpty;
		TaskCondition20307[3]:=((NOT ConveyorIO201081.xEmpty AND ConveyorIO201081.diDesConveyor=20115)
													OR (NOT ConveyorIO20114.xEmpty AND (ConveyorIO20114.diDesConveyor<>20109 OR ConveyorIO20114.diDesConveyor<>20108) ))
													AND ConveyorIo20115.xEmpty;
(*目标地址的传递，横纵分开传递*)
	ConveyorIO20110.diDesConveyorIn:=	ConveyorIO20101.diDesConveyorOut;
	ConveyorIO20111.diDesConveyorIn:=	ConveyorIO20110.diDesConveyorOut;
	ConveyorIO20112.diDesConveyorIn:=	ConveyorIO20111.diDesConveyorOut;
	ConveyorIO20113.diDesConveyorIn:=	ConveyorIO20112.diDesConveyorOut;
	ConveyorIO20114.diDesConveyorIn:=	ConveyorIO20113.diDesConveyorOut;		
(*纵向传递*)
	ConveyorIO20102.diDesConveyorIn:=	ConveyorIO201021.diDesConveyorOut;
	ConveyorIO20103.diDesConveyorIn:=	ConveyorIO201031.diDesConveyorOut;
	ConveyorIO20104.diDesConveyorIn:=	ConveyorIO201041.diDesConveyorOut;
	ConveyorIO20105.diDesConveyorIn:=	ConveyorIO201051.diDesConveyorOut;
	ConveyorIO20106.diDesConveyorIn:=	ConveyorIO201061.diDesConveyorOut;
	ConveyorIO20107.diDesConveyorIn:=	ConveyorIO201071.diDesConveyorOut;
	ConveyorIO20108.diDesConveyorIn:=	ConveyorIO201081.diDesConveyorOut;